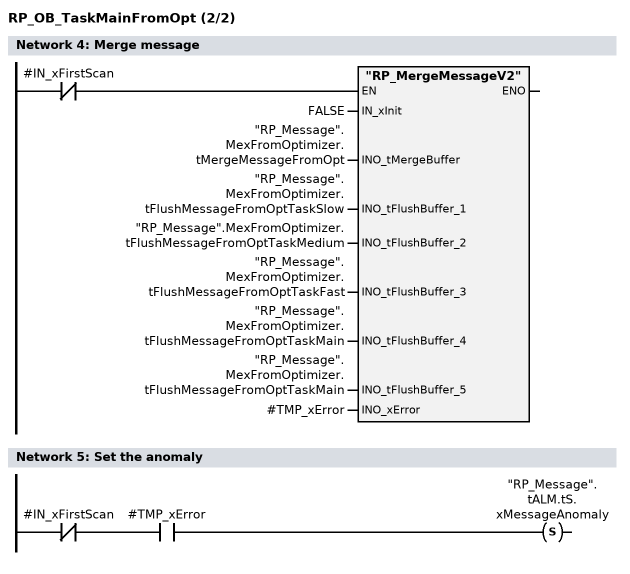
   RUNG wire#powerrail
      I_Contact( #IN_xFirstScan )
      "RP_MergeMessageV2"(IN_xInit := FALSE, INO_tMergeBuffer := "RP_Message".MexFromOptimizer.tMergeMessageFromOpt, INO_tFlushBuffer_1 := "RP_Message".MexFromOptimizer.tFlushMessageFromOptTaskSlow, INO_tFlushBuffer_2 := "RP_Message".MexFromOptimizer.tFlushMessageFromOptTaskMedium, INO_tFlushBuffer_3 := "RP_Message".MexFromOptimizer.tFlushMessageFromOptTaskFast, INO_tFlushBuffer_4 := "RP_Message".MexFromOptimizer.tFlushMessageFromOptTaskMain, INO_tFlushBuffer_5 := "RP_Message".MexFromOptimizer.tFlushMessageFromOptTaskMain, INO_xError := #TMP_xError)
   END_RUNG
   // the same network as SCL:
   IF NOT #IN_xFirstScan THEN
       "RP_MergeMessageV2"(IN_xInit := FALSE,
                           INO_tMergeBuffer := "RP_Message".MexFromOptimizer.tMergeMessageFromOpt,
                           INO_tFlushBuffer_1 := "RP_Message".MexFromOptimizer.tFlushMessageFromOptTaskSlow,
                           INO_tFlushBuffer_2 := "RP_Message".MexFromOptimizer.tFlushMessageFromOptTaskMedium,
                           INO_tFlushBuffer_3 := "RP_Message".MexFromOptimizer.tFlushMessageFromOptTaskFast,
                           INO_tFlushBuffer_4 := "RP_Message".MexFromOptimizer.tFlushMessageFromOptTaskMain,
                           INO_tFlushBuffer_5 := "RP_Message".MexFromOptimizer.tFlushMessageFromOptTaskMain,
                           INO_xError := #TMP_xError);
   END_IF;
END_REGION

REGION Network 5: Set the anomaly
   RUNG wire#powerrail
      I_Contact( #IN_xFirstScan )
      Contact( #TMP_xError )
      S_Coil( "RP_Message".tALM.tS.xMessageAnomaly )
   END_RUNG
   // the same network as SCL:
   IF NOT #IN_xFirstScan AND #TMP_xError THEN "RP_Message".tALM.tS.xMessageAnomaly := TRUE; END_IF;
END_REGION
END_FUNCTION

FUNCTION "RP_AddMessageV2" : Void   // FC27, SCL
TITLE = RP_AddMessage
{ S7_Optimized_Access := 'TRUE' }
AUTHOR : Cigliutt
FAMILY : RP
VERSION : 1.0
// This FC will add one message to the add message buffer
   VAR_INPUT
      IN_xInit : Bool;   // Initialize the buffer container
      IN_dCodeEvent : DInt;   // Event code
      IN_strIndet_Max4Chars : String;   // Station identifier !!! Only 4 char!!!
      IN_dValue1 : DInt;   // Element 1
      IN_dValue2 : DInt;   // Element 2
      IN_dValue3 : DInt;   // Element 3
      IN_dValue4 : DInt;   // Element 4
      IN_dValue5 : DInt;   // Element 5
      IN_dValue6 : DInt;   // Element 6
      IN_dValue7 : DInt;   // Element 7
      IN_dValue8 : DInt;   // Element 8
      IN_dValue9 : DInt;   // Element 9
      IN_dValue10 : DInt;   // Element 10
   END_VAR
   VAR_IN_OUT
      INO_tBuffer : "UDT_RP_AddMessageCont_v2";   // Buffer container
      INO_xError : Bool;   // If =true error on message insert
   END_VAR
   VAR_TEMP
      TMP_dIndex : DInt;
      TMP_dArrayNumEl : DInt;
      TMP_dtDateTime : Date_And_Time;
      TMP_dRetVal : DInt;
   END_VAR
BEGIN
   //Manage the initialization request. Fill to 0 the buffer and the values.
   //After that calculate the space available
   //

   #TMP_dRetVal := RD_LOC_T(#TMP_dtDateTime);

   IF #IN_xInit = true THEN

       //Initialize the values
       #INO_tBuffer.dNumOfMessage := 0;
       #INO_tBuffer.dMaxNumOfMessage := 0;

       //Take the number OF elements OF the array data, reset it AND set the number
       //to iDataMaxElem
       #TMP_dArrayNumEl := "GP_GetArraySize"(INO_vArray := #INO_tBuffer.rgtMessages);

       #INO_tBuffer.dMaxNumOfMessage := #TMP_dArrayNumEl;

       FOR #TMP_dIndex := 0 TO #INO_tBuffer.dMaxNumOfMessage-1 DO
           #INO_tBuffer.rgtMessages[#TMP_dIndex].dCodeEvent := 0;
           #INO_tBuffer.rgtMessages[#TMP_dIndex].strIdent := '';
           #INO_tBuffer.rgtMessages[#TMP_dIndex].dEvent1 := 0;
           #INO_tBuffer.rgtMessages[#TMP_dIndex].dEvent2 := 0;
           #INO_tBuffer.rgtMessages[#TMP_dIndex].dEvent3 := 0;
           #INO_tBuffer.rgtMessages[#TMP_dIndex].dEvent4 := 0;
           #INO_tBuffer.rgtMessages[#TMP_dIndex].dEvent5 := 0;
           #INO_tBuffer.rgtMessages[#TMP_dIndex].dEvent6 := 0;
           #INO_tBuffer.rgtMessages[#TMP_dIndex].dEvent7 := 0;
           #INO_tBuffer.rgtMessages[#TMP_dIndex].dEvent8 := 0;
           #INO_tBuffer.rgtMessages[#TMP_dIndex].dEvent9 := 0;
           #INO_tBuffer.rgtMessages[#TMP_dIndex].dEvent10 := 0;

           #INO_tBuffer.rgtMessages[#TMP_dIndex].dtDateTime := #TMP_dtDateTime;

       END_FOR;


       IF #INO_tBuffer.dMaxNumOfMessage > 0 THEN
           #INO_tBuffer.xInitialized := true;
       END_IF;

       RETURN;
   END_IF;

   //If we are not in initializing mode, copy the input value inside the array.
   //First of all check if the data are consistent
   //
   IF (#INO_tBuffer.xInitialized = false) OR
       (#INO_tBuffer.dMaxNumOfMessage <= 0) OR
       (#INO_tBuffer.dNumOfMessage >=#INO_tBuffer.dMaxNumOfMessage) THEN

       #INO_xError := true;

       RETURN;
   END_IF;

   //Copy the data to the first available index
   //
   #INO_tBuffer.rgtMessages[#INO_tBuffer.dNumOfMessage].dCodeEvent := #IN_dCodeEvent;
   #INO_tBuffer.rgtMessages[#INO_tBuffer.dNumOfMessage].strIdent := #IN_strIndet_Max4Chars;
   #INO_tBuffer.rgtMessages[#INO_tBuffer.dNumOfMessage].dEvent1 := #IN_dValue1;
   #INO_tBuffer.rgtMessages[#INO_tBuffer.dNumOfMessage].dEvent2 := #IN_dValue2;
   #INO_tBuffer.rgtMessages[#INO_tBuffer.dNumOfMessage].dEvent3 := #IN_dValue3;
   #INO_tBuffer.rgtMessages[#INO_tBuffer.dNumOfMessage].dEvent4 := #IN_dValue4;
   #INO_tBuffer.rgtMessages[#INO_tBuffer.dNumOfMessage].dEvent5 := #IN_dValue5;
   #INO_tBuffer.rgtMessages[#INO_tBuffer.dNumOfMessage].dEvent6 := #IN_dValue6;
   #INO_tBuffer.rgtMessages[#INO_tBuffer.dNumOfMessage].dEvent7 := #IN_dValue7;
   #INO_tBuffer.rgtMessages[#INO_tBuffer.dNumOfMessage].dEvent8 := #IN_dValue8;
   #INO_tBuffer.rgtMessages[#INO_tBuffer.dNumOfMessage].dEvent9 := #IN_dValue9;
   #INO_tBuffer.rgtMessages[#INO_tBuffer.dNumOfMessage].dEvent10 := #IN_dValue10;

   #INO_tBuffer.rgtMessages[#INO_tBuffer.dNumOfMessage].dtDateTime := #TMP_dtDateTime;

   //Increment the pointer
   //
   #INO_tBuffer.dNumOfMessage := #INO_tBuffer.dNumOfMessage + 1;
END_FUNCTION

FUNCTION "RP_FlushMessageV2" : Void   // FC39, SCL
TITLE = RP_FlushMessage
{ S7_Optimized_Access := 'TRUE' }
AUTHOR : Cigliutt
FAMILY : RP
VERSION : 1.0
// This FC will flush one AddBuffer to the relative flush buffer
   VAR_INPUT
      IN_xInit : Bool;   // Initialize the buffer container
   END_VAR
   VAR_IN_OUT
      INO_tAddBuffer : "UDT_RP_AddMessageCont_v2";   // Add buffer container
      INO_tFlushBuffer : "UDT_RP_MessageContFlush_v2";   // Flush buffer container
      INO_xError : Bool;   // If =true error on flush
   END_VAR
   VAR_TEMP
      TMP_dIndex : DInt;
      TMP_dArrayNumEl : DInt;
      TMP_dtDateTime : Date_And_Time;
      TMP_dRetVal : DInt;
      TMP_dDataToCopy : DInt;
      TMP_dOldNumMex : DInt;
   END_VAR
BEGIN
   //Manage the initialization request. Fill to 0 the buffer and the values.
   //After that calculate the space available
   //

   #TMP_dRetVal := RD_LOC_T(#TMP_dtDateTime);

   IF #IN_xInit = true THEN

       //Initialize the values
       #INO_tFlushBuffer.dNumOfMessage := 0;
       #INO_tFlushBuffer.dMaxNumOfMessage := 0;

       //Take the number OF elements OF the array data, reset it AND set the number
       //to iDataMaxElem
       #TMP_dArrayNumEl := "GP_GetArraySize"(INO_vArray := #INO_tFlushBuffer.rgtMessages);

       #INO_tFlushBuffer.dMaxNumOfMessage := #TMP_dArrayNumEl;

       //Reset the buffer
       //

       FOR #TMP_dIndex := 0 TO #INO_tFlushBuffer.dMaxNumOfMessage - 1 DO
           #INO_tFlushBuffer.rgtMessages[#TMP_dIndex].dCodeEvent := 0;
           #INO_tFlushBuffer.rgtMessages[#TMP_dIndex].dEvent1 := 0;
           #INO_tFlushBuffer.rgtMessages[#TMP_dIndex].dEvent2 := 0;
           #INO_tFlushBuffer.rgtMessages[#TMP_dIndex].dEvent3 := 0;
           #INO_tFlushBuffer.rgtMessages[#TMP_dIndex].dEvent4 := 0;
           #INO_tFlushBuffer.rgtMessages[#TMP_dIndex].dEvent5 := 0;
           #INO_tFlushBuffer.rgtMessages[#TMP_dIndex].dEvent6 := 0;
           #INO_tFlushBuffer.rgtMessages[#TMP_dIndex].dEvent7 := 0;
           #INO_tFlushBuffer.rgtMessages[#TMP_dIndex].dEvent8 := 0;
           #INO_tFlushBuffer.rgtMessages[#TMP_dIndex].dEvent9 := 0;
           #INO_tFlushBuffer.rgtMessages[#TMP_dIndex].dEvent10 := 0;

           #INO_tFlushBuffer.rgtMessages[#TMP_dIndex].dtDateTime := #TMP_dtDateTime;
           #INO_tFlushBuffer.rgtMessages[#TMP_dIndex].strIdent := '';

       END_FOR;


       IF #INO_tFlushBuffer.dMaxNumOfMessage > 0 THEN
           #INO_tFlushBuffer.xInitialized := true;
       END_IF;

       RETURN;
   END_IF;

   //If we are not in initializing mode, copy the input value inside the array.
   //First of all check if the data are consistent
   //
   IF (#INO_tFlushBuffer.xInitialized = false) OR
       (#INO_tAddBuffer.xInitialized = false) THEN

       #INO_xError := true;

       RETURN;
   END_IF;

   //Check if the flush buffer is free. Otherwise exit
   //
   IF (#INO_tFlushBuffer.dNumOfMessage > 0) THEN
       RETURN;
   END_IF;

   #TMP_dDataToCopy := #INO_tAddBuffer.dNumOfMessage;

   IF (#TMP_dDataToCopy > #INO_tFlushBuffer.dMaxNumOfMessage) THEN
       #TMP_dDataToCopy := #INO_tFlushBuffer.dMaxNumOfMessage;
   END_IF;

   //Copy the data
   #TMP_dRetVal := "GP_BlockMoveStruct"(IN_iSourceIndex := 0,
                        IN_iDestIndex := 0,
                        IN_iCount := DINT_TO_INT(#TMP_dDataToCopy),
                        INO_vSourceArrayStruct := #INO_tAddBuffer.rgtMessages,
                        INO_vDestArrayStruct := #INO_tFlushBuffer.rgtMessages);

   #INO_tFlushBuffer.dNumOfMessage := #TMP_dDataToCopy;

   //Check if some data is remaining. If yes, compact it on the AddBuffer
   //
   IF (#INO_tAddBuffer.dNumOfMessage - #TMP_dDataToCopy) > 0 THEN
       //Copy the data
       #TMP_dRetVal := "GP_BlockMoveStruct"(IN_iSourceIndex := DINT_TO_INT(#INO_tAddBuffer.dNumOfMessage - ( #INO_tAddBuffer.dNumOfMessage - #TMP_dDataToCopy)),
                                            IN_iDestIndex := 0,
                                            IN_iCount := DINT_TO_INT(#INO_tAddBuffer.dNumOfMessage - #TMP_dDataToCopy),
                                            INO_vSourceArrayStruct := #INO_tAddBuffer.rgtMessages,
                                            INO_vDestArrayStruct := #INO_tAddBuffer.rgtMessages);


   END_IF;

   #TMP_dOldNumMex := #INO_tAddBuffer.dNumOfMessage;
   #INO_tAddBuffer.dNumOfMessage := #INO_tAddBuffer.dNumOfMessage - #TMP_dDataToCopy;


   //Data moved, fill the remaining buffer. To increase performance, fill only the data that was used
   //
   FOR #TMP_dIndex := #INO_tAddBuffer.dNumOfMessage TO #TMP_dOldNumMex - 1 DO

       #INO_tAddBuffer.rgtMessages[#TMP_dIndex].dCodeEvent := 0;
       #INO_tAddBuffer.rgtMessages[#TMP_dIndex].dEvent1 := 0;
       #INO_tAddBuffer.rgtMessages[#TMP_dIndex].dEvent2 := 0;
       #INO_tAddBuffer.rgtMessages[#TMP_dIndex].dEvent3 := 0;
       #INO_tAddBuffer.rgtMessages[#TMP_dIndex].dEvent4 := 0;
       #INO_tAddBuffer.rgtMessages[#TMP_dIndex].dEvent5 := 0;
       #INO_tAddBuffer.rgtMessages[#TMP_dIndex].dEvent6 := 0;
       #INO_tAddBuffer.rgtMessages[#TMP_dIndex].dEvent7 := 0;
       #INO_tAddBuffer.rgtMessages[#TMP_dIndex].dEvent8 := 0;
       #INO_tAddBuffer.rgtMessages[#TMP_dIndex].dEvent9 := 0;
       #INO_tAddBuffer.rgtMessages[#TMP_dIndex].dEvent10 := 0;
       #INO_tAddBuffer.rgtMessages[#TMP_dIndex].strIdent := '';

       #INO_tAddBuffer.rgtMessages[#TMP_dIndex].dtDateTime := #TMP_dtDateTime;
   END_FOR;
END_FUNCTION

FUNCTION "RP_MergeMessageV2" : Void   // FC41, SCL
TITLE = RP_MergeMessage
{ S7_Optimized_Access := 'TRUE' }
AUTHOR : Cigliutt
FAMILY : RP
VERSION : 1.0
// This FC will be merge different flush buffer
   VAR_INPUT
      IN_xInit : Bool;   // Initialize the buffer container
   END_VAR
   VAR_IN_OUT
      INO_tMergeBuffer : "UDT_RP_MessageContMerge_v2";   // Merge buffer container
      INO_tFlushBuffer_1 : "UDT_RP_MessageContFlush_v2";   // Flush buffer container #1
      INO_tFlushBuffer_2 : "UDT_RP_MessageContFlush_v2";   // Flush buffer container #2
      INO_tFlushBuffer_3 : "UDT_RP_MessageContFlush_v2";   // Flush buffer container #3
      INO_tFlushBuffer_4 : "UDT_RP_MessageContFlush_v2";   // Flush buffer container #4
      INO_tFlushBuffer_5 : "UDT_RP_MessageContFlush_v2";   // Flush buffer container #5
      INO_xError : Bool;   // If =true error on flush
   END_VAR
   VAR_TEMP
      TMP_dIndex : DInt;
      TMP_dArrayNumEl : DInt;
      TMP_dtDateTime : Date_And_Time;
      TMP_dRetVal : DInt;
      TMP_dDataToCopy : DInt;
      TMP_dOldNumMex : DInt;
      TMP_dActualNumMex : DInt;
   END_VAR
BEGIN
   //Manage the initialization request. Fill to 0 the buffer and the values.
   //After that calculate the space available
   //

   #TMP_dRetVal := RD_LOC_T(#TMP_dtDateTime);
   IF #IN_xInit = true THEN

       //Initialize the values
       #INO_tMergeBuffer.dNumOfMessage := 0;
       #INO_tMergeBuffer.dMaxNumOfMessage := 0;

       //Take the number OF elements OF the array data, reset it AND set the number
       //to iDataMaxElem
       #TMP_dArrayNumEl := "GP_GetArraySize"(INO_vArray := #INO_tMergeBuffer.rgtMessages);

       #INO_tMergeBuffer.dMaxNumOfMessage := #TMP_dArrayNumEl;

       //Reset the buffer
       //

       FOR #TMP_dIndex := 0 TO #INO_tMergeBuffer.dMaxNumOfMessage - 1 DO
           #INO_tMergeBuffer.rgtMessages[#TMP_dIndex].dCodeEvent := 0;
           #INO_tMergeBuffer.rgtMessages[#TMP_dIndex].dEvent1 := 0;
           #INO_tMergeBuffer.rgtMessages[#TMP_dIndex].dEvent2 := 0;
           #INO_tMergeBuffer.rgtMessages[#TMP_dIndex].dEvent3 := 0;
           #INO_tMergeBuffer.rgtMessages[#TMP_dIndex].dEvent4 := 0;
           #INO_tMergeBuffer.rgtMessages[#TMP_dIndex].dEvent5 := 0;
           #INO_tMergeBuffer.rgtMessages[#TMP_dIndex].dEvent6 := 0;
           #INO_tMergeBuffer.rgtMessages[#TMP_dIndex].dEvent7 := 0;
           #INO_tMergeBuffer.rgtMessages[#TMP_dIndex].dEvent8 := 0;
           #INO_tMergeBuffer.rgtMessages[#TMP_dIndex].dEvent9 := 0;
           #INO_tMergeBuffer.rgtMessages[#TMP_dIndex].dEvent10 := 0;
           #INO_tMergeBuffer.rgtMessages[#TMP_dIndex].strIdent := '';

           #INO_tMergeBuffer.rgtMessages[#TMP_dIndex].dtDateTime := #TMP_dtDateTime;

       END_FOR;


       IF #INO_tFlushBuffer_1.dMaxNumOfMessage > 0 THEN
           #INO_tFlushBuffer_1.xInitialized := true;
       END_IF;

       #INO_tMergeBuffer.xInitialized := true;

       RETURN;
   END_IF;

   //If we are not in initializing mode, copy the input value inside the array.
   //First of all check if the data are consistent
   //
   IF (#INO_tMergeBuffer.xInitialized = false) OR
       (#INO_tFlushBuffer_1.xInitialized = false) OR
       (#INO_tFlushBuffer_2.xInitialized = false) OR
       (#INO_tFlushBuffer_3.xInitialized = false) OR
       (#INO_tFlushBuffer_4.xInitialized = false) OR
       (#INO_tFlushBuffer_5.xInitialized = false) THEN

       #INO_xError := true;

       RETURN;
   END_IF;

   //Check if the merge buffer is free. Otherwise exit
   //
   IF (#INO_tMergeBuffer.dNumOfMessage > 0) THEN
       RETURN;
   END_IF;


   ///*********************************** FLUSH BUFFER #1

   //Check if the first flush buffer, has data inside
   IF (#INO_tFlushBuffer_1.dNumOfMessage > 0) THEN

       #TMP_dDataToCopy := #INO_tFlushBuffer_1.dNumOfMessage;

       IF (#TMP_dDataToCopy > #INO_tMergeBuffer.dMaxNumOfMessage) THEN
           #TMP_dDataToCopy := #INO_tMergeBuffer.dMaxNumOfMessage;
       END_IF;

       //Copy the data
       #TMP_dRetVal := "GP_BlockMoveStruct"(IN_iSourceIndex := 0,
                                            IN_iDestIndex := 0,
                                            IN_iCount := DINT_TO_INT(#TMP_dDataToCopy),
                                            INO_vSourceArrayStruct := #INO_tFlushBuffer_1.rgtMessages,
                                            INO_vDestArrayStruct := #INO_tMergeBuffer.rgtMessages);

       #INO_tMergeBuffer.dNumOfMessage := #TMP_dDataToCopy;

       //Check if some data is remaining. If yes, compact it on the FlushBuffer
       //
       IF (#INO_tFlushBuffer_1.dNumOfMessage - #TMP_dDataToCopy) > 0 THEN
           //Copy the data
           #TMP_dRetVal := "GP_BlockMoveStruct"(IN_iSourceIndex := DINT_TO_INT(#INO_tFlushBuffer_1.dNumOfMessage - (#INO_tFlushBuffer_1.dNumOfMessage - #TMP_dDataToCopy)),
                                                IN_iDestIndex := 0,
                                                IN_iCount := DINT_TO_INT(#INO_tFlushBuffer_1.dNumOfMessage - #TMP_dDataToCopy),
                                                INO_vSourceArrayStruct := #INO_tFlushBuffer_1.rgtMessages,
                                                INO_vDestArrayStruct := #INO_tFlushBuffer_1.rgtMessages);


       END_IF;

       #TMP_dOldNumMex := #INO_tFlushBuffer_1.dNumOfMessage;
       #TMP_dActualNumMex := #INO_tFlushBuffer_1.dNumOfMessage - #TMP_dDataToCopy;


       //Data moved, fill the remaining buffer. To increase performance, fill only the data that was used
       //
       FOR #TMP_dIndex := #TMP_dActualNumMex TO #TMP_dOldNumMex - 1 DO

           #INO_tFlushBuffer_1.rgtMessages[#TMP_dIndex].dCodeEvent := 0;
           #INO_tFlushBuffer_1.rgtMessages[#TMP_dIndex].dEvent1 := 0;
           #INO_tFlushBuffer_1.rgtMessages[#TMP_dIndex].dEvent2 := 0;
           #INO_tFlushBuffer_1.rgtMessages[#TMP_dIndex].dEvent3 := 0;
           #INO_tFlushBuffer_1.rgtMessages[#TMP_dIndex].dEvent4 := 0;
           #INO_tFlushBuffer_1.rgtMessages[#TMP_dIndex].dEvent5 := 0;
           #INO_tFlushBuffer_1.rgtMessages[#TMP_dIndex].dEvent6 := 0;
           #INO_tFlushBuffer_1.rgtMessages[#TMP_dIndex].dEvent7 := 0;
           #INO_tFlushBuffer_1.rgtMessages[#TMP_dIndex].dEvent8 := 0;
           #INO_tFlushBuffer_1.rgtMessages[#TMP_dIndex].dEvent9 := 0;
           #INO_tFlushBuffer_1.rgtMessages[#TMP_dIndex].dEvent10 := 0;
           #INO_tFlushBuffer_1.rgtMessages[#TMP_dIndex].strIdent := '';

           #INO_tFlushBuffer_1.rgtMessages[#TMP_dIndex].dtDateTime := #TMP_dtDateTime;
       END_FOR;

       #INO_tFlushBuffer_1.dNumOfMessage := #TMP_dActualNumMex;

   END_IF;

   //RETURN;
   ///*********************************** FLUSH BUFFER #2

   //Check if the first flush buffer, has data inside
   IF (#INO_tFlushBuffer_2.dNumOfMessage > 0) AND (#INO_tMergeBuffer.dNumOfMessage < #INO_tMergeBuffer.dMaxNumOfMessage) THEN

       #TMP_dDataToCopy := #INO_tFlushBuffer_2.dNumOfMessage;

       IF (#TMP_dDataToCopy + #INO_tMergeBuffer.dNumOfMessage > #INO_tMergeBuffer.dMaxNumOfMessage) THEN
           #TMP_dDataToCopy := #INO_tMergeBuffer.dMaxNumOfMessage - #INO_tMergeBuffer.dNumOfMessage;
       END_IF;

       //Copy the data
       #TMP_dRetVal := "GP_BlockMoveStruct"(IN_iSourceIndex := 0,
                                            IN_iDestIndex := DINT_TO_INT(#INO_tMergeBuffer.dNumOfMessage),
                                            IN_iCount := DINT_TO_INT(#TMP_dDataToCopy),
                                            INO_vSourceArrayStruct := #INO_tFlushBuffer_2.rgtMessages,
                                            INO_vDestArrayStruct := #INO_tMergeBuffer.rgtMessages);

       #INO_tMergeBuffer.dNumOfMessage := #INO_tMergeBuffer.dNumOfMessage + #TMP_dDataToCopy;

       //Check if some data is remaining. If yes, compact it on the FlushBuffer
       //
       IF (#INO_tFlushBuffer_2.dNumOfMessage - #TMP_dDataToCopy) > 0 THEN
           //Copy the data
           #TMP_dRetVal := "GP_BlockMoveStruct"(IN_iSourceIndex := DINT_TO_INT(#INO_tFlushBuffer_2.dNumOfMessage - (#INO_tFlushBuffer_2.dNumOfMessage - #TMP_dDataToCopy)),
                                                IN_iDestIndex := 0,
                                                IN_iCount := DINT_TO_INT(#INO_tFlushBuffer_2.dNumOfMessage - #TMP_dDataToCopy),
                                                INO_vSourceArrayStruct := #INO_tFlushBuffer_2.rgtMessages,
                                                INO_vDestArrayStruct := #INO_tFlushBuffer_2.rgtMessages);


       END_IF;

       #TMP_dOldNumMex := #INO_tFlushBuffer_2.dNumOfMessage;
       #TMP_dActualNumMex := #INO_tFlushBuffer_2.dNumOfMessage - #TMP_dDataToCopy;



       //Data moved, fill the remaining buffer. To increase performance, fill only the data that was used
       //
       FOR #TMP_dIndex := #TMP_dActualNumMex TO #TMP_dOldNumMex - 1 DO

           #INO_tFlushBuffer_2.rgtMessages[#TMP_dIndex].dCodeEvent := 0;
           #INO_tFlushBuffer_2.rgtMessages[#TMP_dIndex].dEvent1 := 0;
           #INO_tFlushBuffer_2.rgtMessages[#TMP_dIndex].dEvent2 := 0;
           #INO_tFlushBuffer_2.rgtMessages[#TMP_dIndex].dEvent3 := 0;
           #INO_tFlushBuffer_2.rgtMessages[#TMP_dIndex].dEvent4 := 0;
           #INO_tFlushBuffer_2.rgtMessages[#TMP_dIndex].dEvent5 := 0;
           #INO_tFlushBuffer_2.rgtMessages[#TMP_dIndex].dEvent6 := 0;
           #INO_tFlushBuffer_2.rgtMessages[#TMP_dIndex].dEvent7 := 0;
           #INO_tFlushBuffer_2.rgtMessages[#TMP_dIndex].dEvent8 := 0;
           #INO_tFlushBuffer_2.rgtMessages[#TMP_dIndex].dEvent9 := 0;
           #INO_tFlushBuffer_2.rgtMessages[#TMP_dIndex].dEvent10 := 0;

           #INO_tFlushBuffer_2.rgtMessages[#TMP_dIndex].strIdent := '';
           #INO_tFlushBuffer_2.rgtMessages[#TMP_dIndex].dtDateTime := #TMP_dtDateTime;
       END_FOR;

       #INO_tFlushBuffer_2.dNumOfMessage := #TMP_dActualNumMex;
   END_IF;


   ///*********************************** FLUSH BUFFER #3


   //Check if the first flush buffer, has data inside
   IF (#INO_tFlushBuffer_3.dNumOfMessage > 0) AND (#INO_tMergeBuffer.dNumOfMessage < #INO_tMergeBuffer.dMaxNumOfMessage) THEN

       #TMP_dDataToCopy := #INO_tFlushBuffer_3.dNumOfMessage;

       IF (#TMP_dDataToCopy + #INO_tMergeBuffer.dNumOfMessage > #INO_tMergeBuffer.dMaxNumOfMessage) THEN
           #TMP_dDataToCopy := #INO_tMergeBuffer.dMaxNumOfMessage - #INO_tMergeBuffer.dNumOfMessage;
       END_IF;

       //Copy the data
       #TMP_dRetVal := "GP_BlockMoveStruct"(IN_iSourceIndex := 0,
                                            IN_iDestIndex := DINT_TO_INT(#INO_tMergeBuffer.dNumOfMessage),
                                            IN_iCount := DINT_TO_INT(#TMP_dDataToCopy),
                                            INO_vSourceArrayStruct := #INO_tFlushBuffer_3.rgtMessages,
                                            INO_vDestArrayStruct := #INO_tMergeBuffer.rgtMessages);

       #INO_tMergeBuffer.dNumOfMessage := #INO_tMergeBuffer.dNumOfMessage + #TMP_dDataToCopy;

       //Check if some data is remaining. If yes, compact it on the FlushBuffer
       //
       IF (#INO_tFlushBuffer_3.dNumOfMessage - #TMP_dDataToCopy) > 0 THEN
           //Copy the data
           #TMP_dRetVal := "GP_BlockMoveStruct"(IN_iSourceIndex := DINT_TO_INT(#INO_tFlushBuffer_3.dNumOfMessage - (#INO_tFlushBuffer_3.dNumOfMessage - #TMP_dDataToCopy)),
                                                IN_iDestIndex := 0,
                                                IN_iCount := DINT_TO_INT(#INO_tFlushBuffer_3.dNumOfMessage - #TMP_dDataToCopy),
                                                INO_vSourceArrayStruct := #INO_tFlushBuffer_3.rgtMessages,
                                                INO_vDestArrayStruct := #INO_tFlushBuffer_3.rgtMessages);


       END_IF;

       #TMP_dOldNumMex := #INO_tFlushBuffer_3.dNumOfMessage;
       #TMP_dActualNumMex := #INO_tFlushBuffer_3.dNumOfMessage - #TMP_dDataToCopy;


       //Data moved, fill the remaining buffer. To increase performance, fill only the data that was used
       //
       FOR #TMP_dIndex := #TMP_dActualNumMex TO #TMP_dOldNumMex - 1 DO

           #INO_tFlushBuffer_3.rgtMessages[#TMP_dIndex].dCodeEvent := 0;
           #INO_tFlushBuffer_3.rgtMessages[#TMP_dIndex].dEvent1 := 0;
           #INO_tFlushBuffer_3.rgtMessages[#TMP_dIndex].dEvent2 := 0;
           #INO_tFlushBuffer_3.rgtMessages[#TMP_dIndex].dEvent3 := 0;
           #INO_tFlushBuffer_3.rgtMessages[#TMP_dIndex].dEvent4 := 0;
           #INO_tFlushBuffer_3.rgtMessages[#TMP_dIndex].dEvent5 := 0;
           #INO_tFlushBuffer_3.rgtMessages[#TMP_dIndex].dEvent6 := 0;
           #INO_tFlushBuffer_3.rgtMessages[#TMP_dIndex].dEvent7 := 0;
           #INO_tFlushBuffer_3.rgtMessages[#TMP_dIndex].dEvent8 := 0;
           #INO_tFlushBuffer_3.rgtMessages[#TMP_dIndex].dEvent9 := 0;
           #INO_tFlushBuffer_3.rgtMessages[#TMP_dIndex].dEvent10 := 0;
           #INO_tFlushBuffer_3.rgtMessages[#TMP_dIndex].strIdent := '';

           #INO_tFlushBuffer_3.rgtMessages[#TMP_dIndex].dtDateTime := #TMP_dtDateTime;
       END_FOR;

       #INO_tFlushBuffer_3.dNumOfMessage := #TMP_dActualNumMex;


   END_IF;


   ///*********************************** FLUSH BUFFER #4


   //Check if the first flush buffer, has data inside
   IF (#INO_tFlushBuffer_4.dNumOfMessage > 0) AND (#INO_tMergeBuffer.dNumOfMessage < #INO_tMergeBuffer.dMaxNumOfMessage) THEN

       #TMP_dDataToCopy := #INO_tFlushBuffer_4.dNumOfMessage;

       IF (#TMP_dDataToCopy + #INO_tMergeBuffer.dNumOfMessage > #INO_tMergeBuffer.dMaxNumOfMessage) THEN
           #TMP_dDataToCopy := #INO_tMergeBuffer.dMaxNumOfMessage - #INO_tMergeBuffer.dNumOfMessage;
       END_IF;

       //Copy the data
       #TMP_dRetVal := "GP_BlockMoveStruct"(IN_iSourceIndex := 0,
                                            IN_iDestIndex := DINT_TO_INT(#INO_tMergeBuffer.dNumOfMessage),
                                            IN_iCount := DINT_TO_INT(#TMP_dDataToCopy),
                                            INO_vSourceArrayStruct := #INO_tFlushBuffer_4.rgtMessages,
                                            INO_vDestArrayStruct := #INO_tMergeBuffer.rgtMessages);

       #INO_tMergeBuffer.dNumOfMessage := #INO_tMergeBuffer.dNumOfMessage + #TMP_dDataToCopy;

       //Check if some data is remaining. If yes, compact it on the FlushBuffer
       //
       IF (#INO_tFlushBuffer_4.dNumOfMessage - #TMP_dDataToCopy) > 0 THEN
           //Copy the data
           #TMP_dRetVal := "GP_BlockMoveStruct"(IN_iSourceIndex := DINT_TO_INT(#INO_tFlushBuffer_4.dNumOfMessage - (#INO_tFlushBuffer_4.dNumOfMessage - #TMP_dDataToCopy)),
                                                IN_iDestIndex := 0,
                                                IN_iCount := DINT_TO_INT(#INO_tFlushBuffer_4.dNumOfMessage - #TMP_dDataToCopy),
                                                INO_vSourceArrayStruct := #INO_tFlushBuffer_4.rgtMessages,
                                                INO_vDestArrayStruct := #INO_tFlushBuffer_4.rgtMessages);


       END_IF;

       #TMP_dOldNumMex := #INO_tFlushBuffer_4.dNumOfMessage;
       #TMP_dActualNumMex := #INO_tFlushBuffer_4.dNumOfMessage - #TMP_dDataToCopy;


       //Data moved, fill the remaining buffer. To increase performance, fill only the data that was used
       //
       FOR #TMP_dIndex := #TMP_dActualNumMex TO #TMP_dOldNumMex - 1 DO

           #INO_tFlushBuffer_4.rgtMessages[#TMP_dIndex].dCodeEvent := 0;
           #INO_tFlushBuffer_4.rgtMessages[#TMP_dIndex].dEvent1 := 0;
           #INO_tFlushBuffer_4.rgtMessages[#TMP_dIndex].dEvent2 := 0;
           #INO_tFlushBuffer_4.rgtMessages[#TMP_dIndex].dEvent3 := 0;
           #INO_tFlushBuffer_4.rgtMessages[#TMP_dIndex].dEvent4 := 0;
           #INO_tFlushBuffer_4.rgtMessages[#TMP_dIndex].dEvent5 := 0;
           #INO_tFlushBuffer_4.rgtMessages[#TMP_dIndex].dEvent6 := 0;
           #INO_tFlushBuffer_4.rgtMessages[#TMP_dIndex].dEvent7 := 0;
           #INO_tFlushBuffer_4.rgtMessages[#TMP_dIndex].dEvent8 := 0;
           #INO_tFlushBuffer_4.rgtMessages[#TMP_dIndex].dEvent9 := 0;
           #INO_tFlushBuffer_4.rgtMessages[#TMP_dIndex].dEvent10 := 0;
           #INO_tFlushBuffer_4.rgtMessages[#TMP_dIndex].strIdent := '';

           #INO_tFlushBuffer_4.rgtMessages[#TMP_dIndex].dtDateTime := #TMP_dtDateTime;
       END_FOR;

       #INO_tFlushBuffer_4.dNumOfMessage := #TMP_dActualNumMex;


   END_IF;


   ///*********************************** FLUSH BUFFER #5


   //Check if the first flush buffer, has data inside
   IF (#INO_tFlushBuffer_5.dNumOfMessage > 0) AND (#INO_tMergeBuffer.dNumOfMessage < #INO_tMergeBuffer.dMaxNumOfMessage) THEN

       #TMP_dDataToCopy := #INO_tFlushBuffer_5.dNumOfMessage;

       IF (#TMP_dDataToCopy + #INO_tMergeBuffer.dNumOfMessage > #INO_tMergeBuffer.dMaxNumOfMessage) THEN
           #TMP_dDataToCopy := #INO_tMergeBuffer.dMaxNumOfMessage - #INO_tMergeBuffer.dNumOfMessage;
       END_IF;

       //Copy the data
       #TMP_dRetVal := "GP_BlockMoveStruct"(IN_iSourceIndex := 0,
                                            IN_iDestIndex := DINT_TO_INT(#INO_tMergeBuffer.dNumOfMessage),
                                            IN_iCount := DINT_TO_INT(#TMP_dDataToCopy),
                                            INO_vSourceArrayStruct := #INO_tFlushBuffer_5.rgtMessages,
                                            INO_vDestArrayStruct := #INO_tMergeBuffer.rgtMessages);

       #INO_tMergeBuffer.dNumOfMessage := #INO_tMergeBuffer.dNumOfMessage + #TMP_dDataToCopy;

       //Check if some data is remaining. If yes, compact it on the FlushBuffer
       //
       IF (#INO_tFlushBuffer_5.dNumOfMessage - #TMP_dDataToCopy) > 0 THEN
           //Copy the data
           #TMP_dRetVal := "GP_BlockMoveStruct"(IN_iSourceIndex := DINT_TO_INT(#INO_tFlushBuffer_5.dNumOfMessage - (#INO_tFlushBuffer_5.dNumOfMessage - #TMP_dDataToCopy)),
                                                IN_iDestIndex := 0,
                                                IN_iCount := DINT_TO_INT(#INO_tFlushBuffer_5.dNumOfMessage - #TMP_dDataToCopy),
                                                INO_vSourceArrayStruct := #INO_tFlushBuffer_5.rgtMessages,
                                                INO_vDestArrayStruct := #INO_tFlushBuffer_5.rgtMessages);


       END_IF;

       #TMP_dOldNumMex := #INO_tFlushBuffer_5.dNumOfMessage;
       #TMP_dActualNumMex := #INO_tFlushBuffer_5.dNumOfMessage - #TMP_dDataToCopy;

       //Data moved, fill the remaining buffer. To increase performance, fill only the data that was used
       //
       FOR #TMP_dIndex := #TMP_dActualNumMex TO #TMP_dOldNumMex - 1 DO

           #INO_tFlushBuffer_5.rgtMessages[#TMP_dIndex].dCodeEvent := 0;
           #INO_tFlushBuffer_5.rgtMessages[#TMP_dIndex].dEvent1 := 0;
           #INO_tFlushBuffer_5.rgtMessages[#TMP_dIndex].dEvent2 := 0;
           #INO_tFlushBuffer_5.rgtMessages[#TMP_dIndex].dEvent3 := 0;
           #INO_tFlushBuffer_5.rgtMessages[#TMP_dIndex].dEvent4 := 0;
           #INO_tFlushBuffer_5.rgtMessages[#TMP_dIndex].dEvent5 := 0;
           #INO_tFlushBuffer_5.rgtMessages[#TMP_dIndex].dEvent6 := 0;
           #INO_tFlushBuffer_5.rgtMessages[#TMP_dIndex].dEvent7 := 0;
           #INO_tFlushBuffer_5.rgtMessages[#TMP_dIndex].dEvent8 := 0;
           #INO_tFlushBuffer_5.rgtMessages[#TMP_dIndex].dEvent9 := 0;
           #INO_tFlushBuffer_5.rgtMessages[#TMP_dIndex].dEvent10 := 0;

           #INO_tFlushBuffer_5.rgtMessages[#TMP_dIndex].dtDateTime := #TMP_dtDateTime;
           #INO_tFlushBuffer_5.rgtMessages[#TMP_dIndex].strIdent := '';
       END_FOR;

       #INO_tFlushBuffer_5.dNumOfMessage := #TMP_dActualNumMex;


   END_IF;

   //Clear the remaining data
   FOR #TMP_dIndex := #INO_tMergeBuffer.dNumOfMessage TO #INO_tMergeBuffer.dMaxNumOfMessage - 1 DO

           #INO_tMergeBuffer.rgtMessages[#TMP_dIndex].dCodeEvent := 0;
           #INO_tMergeBuffer.rgtMessages[#TMP_dIndex].dEvent1 := 0;
           #INO_tMergeBuffer.rgtMessages[#TMP_dIndex].dEvent2 := 0;
           #INO_tMergeBuffer.rgtMessages[#TMP_dIndex].dEvent3 := 0;
           #INO_tMergeBuffer.rgtMessages[#TMP_dIndex].dEvent4 := 0;
           #INO_tMergeBuffer.rgtMessages[#TMP_dIndex].dEvent5 := 0;
           #INO_tMergeBuffer.rgtMessages[#TMP_dIndex].dEvent6 := 0;
           #INO_tMergeBuffer.rgtMessages[#TMP_dIndex].dEvent7 := 0;
           #INO_tMergeBuffer.rgtMessages[#TMP_dIndex].dEvent8 := 0;
           #INO_tMergeBuffer.rgtMessages[#TMP_dIndex].dEvent9 := 0;
           #INO_tMergeBuffer.rgtMessages[#TMP_dIndex].dEvent10 := 0;
           #INO_tMergeBuffer.rgtMessages[#TMP_dIndex].strIdent := '';
           #INO_tMergeBuffer.rgtMessages[#TMP_dIndex].dtDateTime := #TMP_dtDateTime;

   END_FOR;
END_FUNCTION

FUNCTION "RP_ExtractMessageV2" : Void   // FC42, SCL
TITLE = RP_ExtractMessage
{ S7_Optimized_Access := 'TRUE' }
AUTHOR : Cigliutt
FAMILY : RP
VERSION : 1.01
// This FC will extract each call one message from the merge buffer
   VAR_OUTPUT
      OUT_xDataAvailable : Bool;   // If true data available to read
      OUT_dCodeEvent : DInt;   // Event code
      OUT_dtDateTime : Date_And_Time;   // Event date and time
      OUT_strIdent : String;
      OUT_dValue1 : DInt;   // Event value 1
      OUT_dValue2 : DInt;   // Event value 2
      OUT_dValue3 : DInt;   // Event value 3
      OUT_dValue4 : DInt;   // Event value 4
      OUT_dValue5 : DInt;   // Event value 5
      OUT_dValue6 : DInt;   // Event value 6
      OUT_dValue7 : DInt;   // Event value 7
      OUT_dValue8 : DInt;   // Event value 8
      OUT_dValue9 : DInt;   // Event value 9
      OUT_dValue10 : DInt;   // Event value 10
   END_VAR
   VAR_IN_OUT
      INO_tMergeBuffer : "UDT_RP_MessageContMerge_v2";   // Merge buffer container
      INO_xError : Bool;   // If =true error on buffer
   END_VAR
   VAR_TEMP
      TMP_dIndex : DInt;
      TMP_dArrayNumEl : DInt;
      TMP_dtDateTime : Date_And_Time;
      TMP_dRetVal : DInt;
   END_VAR
BEGIN
   //Check if the buffer is initialized, otherwise exit
   //
   #OUT_xDataAvailable := false;

   IF #INO_tMergeBuffer.xInitialized = false THEN

       #INO_xError := true;

       RETURN;
   END_IF;

   //Check if data are available
   IF (#INO_tMergeBuffer.dNumOfMessage > 0) THEN


   //Take the first message, and copy to the out
   //

       #OUT_dCodeEvent := #INO_tMergeBuffer.rgtMessages[0].dCodeEvent;
       #OUT_dtDateTime := #INO_tMergeBuffer.rgtMessages[0].dtDateTime;
       #OUT_strIdent := #INO_tMergeBuffer.rgtMessages[0].strIdent;
       #OUT_dValue1 := #INO_tMergeBuffer.rgtMessages[0].dEvent1;
       #OUT_dValue2 := #INO_tMergeBuffer.rgtMessages[0].dEvent2;
       #OUT_dValue3 := #INO_tMergeBuffer.rgtMessages[0].dEvent3;
       #OUT_dValue4 := #INO_tMergeBuffer.rgtMessages[0].dEvent4;
       #OUT_dValue5 := #INO_tMergeBuffer.rgtMessages[0].dEvent5;
       #OUT_dValue6 := #INO_tMergeBuffer.rgtMessages[0].dEvent6;
       #OUT_dValue7 := #INO_tMergeBuffer.rgtMessages[0].dEvent7;
       #OUT_dValue8 := #INO_tMergeBuffer.rgtMessages[0].dEvent8;
       #OUT_dValue9 := #INO_tMergeBuffer.rgtMessages[0].dEvent9;
       #OUT_dValue10 := #INO_tMergeBuffer.rgtMessages[0].dEvent10;



   //Fill to 0 the read data
   //
       #INO_tMergeBuffer.rgtMessages[0].dCodeEvent := 0;
       #INO_tMergeBuffer.rgtMessages[0].strIdent := '';
       #INO_tMergeBuffer.rgtMessages[0].dEvent1 := 0;
       #INO_tMergeBuffer.rgtMessages[0].dEvent2 := 0;
       #INO_tMergeBuffer.rgtMessages[0].dEvent3 := 0;
       #INO_tMergeBuffer.rgtMessages[0].dEvent4 := 0;
       #INO_tMergeBuffer.rgtMessages[0].dEvent5 := 0;
       #INO_tMergeBuffer.rgtMessages[0].dEvent6 := 0;
       #INO_tMergeBuffer.rgtMessages[0].dEvent7 := 0;
       #INO_tMergeBuffer.rgtMessages[0].dEvent8 := 0;
       #INO_tMergeBuffer.rgtMessages[0].dEvent9 := 0;
       #INO_tMergeBuffer.rgtMessages[0].dEvent10 := 0;

       IF (#INO_tMergeBuffer.dNumOfMessage = 1) THEN
           #INO_tMergeBuffer.dNumOfMessage := 0;
       ELSE
           //Compact the array    
           #TMP_dRetVal := "GP_BlockMoveStruct"(IN_iSourceIndex := 1,
                                IN_iDestIndex := 0,
                                IN_iCount := DINT_TO_INT(#INO_tMergeBuffer.dNumOfMessage - 1),
                                INO_vSourceArrayStruct := #INO_tMergeBuffer.rgtMessages,
                                INO_vDestArrayStruct := #INO_tMergeBuffer.rgtMessages);